(*ConveyorIO70150.xPosLimit:=X49;*)						
ConveyorIO70150.xCWPresent:=X48;						
Y248:=ConveyorIO70150.xMotorCW;						
ConveyorIO70150.xForward:=M564;						
M350:= NOT ConveyorIO70150.xEmpty;						
M749:=ConveyorIO70150.xError;						
ConveyorIO70150.diDeviceID:=70150;						

ConveyorIO70151.xPosLimit:=X4B;						
ConveyorIO70151.xCWPresent:=X4A;						
Y249:=ConveyorIO70151.xMotorCCW;						
ConveyorIO70151.xBackward:=M565;						
M351:= NOT ConveyorIO70151.xEmpty;						
M750:=ConveyorIO70151.xError;						
ConveyorIO70151.diDeviceID:=70151;						

ConveyorIO70152.xCWPresent:=X4D;						
Y24A:=ConveyorIO70152.xMotorCW;						
ConveyorIO70152.xForward:=M566;						
M352:= NOT ConveyorIO70152.xEmpty;						
M751:=ConveyorIO70152.xError;						
ConveyorIO70152.diDeviceID:=70152;			
ConveyorIO70152.tLoadDelay:=T#7S;			

ConveyorIO70153.xCWPresent:=X4D;						
Y24B:=ConveyorIO70153.xMotorCW;						
ConveyorIO70153.xForward:=M567;						
M353:= NOT ConveyorIO70153.xEmpty;						
M752:=ConveyorIO70153.xError;						
ConveyorIO70153.diDeviceID:=70153;						

ConveyorIO70154.xPosLimit:=X4F;						
ConveyorIO70154.xCWPresent:=X4E;						
Y24C:=ConveyorIO70154.xMotorCW;						
ConveyorIO70154.xForward:=M568;						
M354:= NOT ConveyorIO70154.xEmpty;						
M753:=ConveyorIO70154.xError;						
ConveyorIO70154.diDeviceID:=70154;		
ConveyorIO70154.tLoadDelay:=T#4S;				
				
ConveyorIO70155.xCWPresent:=X50;						
Y24D:=ConveyorIO70155.xMotorCW;						
ConveyorIO70155.xBackward:=M569;						
M355:= NOT ConveyorIO70155.xEmpty;						
M754:=ConveyorIO70155.xError;						
ConveyorIO70155.diDeviceID:=70155;		
ConveyorIO70155.tLoadDelay:=T#4S;						

ConveyorIO70156.xPosLimit:=NOT  X53;						
ConveyorIO70156.xCWPresent:=X52;						
Y24E:=ConveyorIO70156.xMotorCW;						
ConveyorIO70156.xForward:=M570;						
M356:= NOT ConveyorIO70156.xEmpty;						
M755:=ConveyorIO70156.xError;						
ConveyorIO70156.diDeviceID:=70156;						

ConveyorIO70157.xCWPresent:=X54;						
Y24F:=ConveyorIO70157.xMotorCW;						
ConveyorIO70157.xForward:=M571;						
M357:= NOT ConveyorIO70157.xEmpty;						
M756:=ConveyorIO70157.xError;						
ConveyorIO70157.diDeviceID:=70157;						

ConveyorIO70158.xPosLimit:=X56;						
ConveyorIO70158.xCWPresent:=X55;						
Y250:=ConveyorIO70158.xMotorCW;						
ConveyorIO70158.xForward:=M572;						
M358:= NOT ConveyorIO70158.xEmpty;						
M757:=ConveyorIO70158.xError;						
ConveyorIO70158.diDeviceID:=70158;						

(*ConveyorIO70159.xPosLimit:=X57;	*)					
ConveyorIO70159.xCWPresent:=X57;						
Y251:=ConveyorIO70159.xMotorCW;						
ConveyorIO70159.xBackward:=M573;						
M359:= NOT ConveyorIO70159.xEmpty;						
M758:=ConveyorIO70159.xError;						
ConveyorIO70159.diDeviceID:=70159;						

ConveyorIO70160.xCWPresent:=X59;						
Y252:=ConveyorIO70160.xMotorCW;						
ConveyorIO70160.xForward:=M574;						
M360:= NOT ConveyorIO70160.xEmpty;						
M759:=ConveyorIO70160.xError;						
ConveyorIO70160.diDeviceID:=70160;		
ConveyorIO70160.tLoadDelay:=T#7S;				

ConveyorIO70161.xCWPresent:=X5A;						
Y253:=ConveyorIO70161.xMotorCW;						
ConveyorIO70161.xForward:=M575;						
M361:= NOT ConveyorIO70161.xEmpty;						
M760:=ConveyorIO70161.xError;						
ConveyorIO70161.diDeviceID:=70161;						

(*ConveyorIO70162.xPosLimit:=X5C;	*)					
ConveyorIO70162.xCWPresent:=X5B;						
Y254:=ConveyorIO70162.xMotorCW;						
ConveyorIO70162.xForward:=M576;						
M362:= NOT ConveyorIO70162.xEmpty;						
M761:=ConveyorIO70162.xError;						
ConveyorIO70162.diDeviceID:=70162;						
ConveyorIO70162.tLoadDelay:=T#5S;

(*ConveyorIO70163.xPosLimit:=X5E;	*)					
ConveyorIO70163.xCWPresent:=X5D;						
Y305:=ConveyorIO70163.xMotorCW ;						
ConveyorIO70163.xBackward:=M577;						
M363:= NOT ConveyorIO70163.xEmpty;						
M762:=ConveyorIO70163.xError;						
ConveyorIO70163.diDeviceID:=70163;	
ConveyorIO70163.tLoadDelay:=t#4s;

ConveyorIO70164.xCWPresent:=X5F;						
Y256:=ConveyorIO70164.xMotorCW OR M800;						
ConveyorIO70164.xForward:=M578;						
M364:= NOT ConveyorIO70164.xEmpty;						
M763:=ConveyorIO70164.xError;						
ConveyorIO70164.diDeviceID:=70164;			
ConveyorIO70164.tLoadDelay:=T#4s;			

ConveyorIO70165.xCWPresent:=X61;						
Y257:=ConveyorIO70165.xMotorCW OR ConveyorIO70165_2.xMotorCW;						
ConveyorIO70165.xForward:=M579;						
M365:= NOT ConveyorIO70165.xEmpty;						
M764:=ConveyorIO70165.xError;						
ConveyorIO70165.diDeviceID:=70165;		
ConveyorIO70165.tLoadDelay:=T#4200MS;


ConveyorIO70165_1.xCWPresent:=	X5F;
ConveyorIO70165_1.diDeviceID:=70164;		

ConveyorIO70165_2.xCWPresent:=	X60;
ConveyorIO70165_2.diDeviceID:=70165;		
ConveyorIO70165_2.tLoadDelay:=T#4500MS;

ConveyorIO70166.xCWPresent:=X62;						
Y258:=ConveyorIO70166.xMotorCW;						
ConveyorIO70166.xForward:=M580;						
M366:= NOT ConveyorIO70166.xEmpty;						
M765:=ConveyorIO70166.xError;						
ConveyorIO70166.diDeviceID:=70166;						
ConveyorIO70166.tLoadDelay:=T#6S;

ConveyorIO70167.xCWPresent:=X63;						
Y259:=ConveyorIO70167.xMotorCW;						
ConveyorIO70167.xForward:=M581;						
M367:= NOT ConveyorIO70167.xEmpty;						
M766:=ConveyorIO70167.xError;						
ConveyorIO70167.diDeviceID:=70167;		
ConveyorIO70167.tLoadDelay:=T#8S;				

ConveyorIO70168.xCWPresent:=X65;						
Y25A:=ConveyorIO70168.xMotorCW OR ConveyorIO70168_1.xMotorCW;						
ConveyorIO70168.xForward:=M582;						
M368:= NOT ConveyorIO70168.xEmpty;						
M767:=ConveyorIO70168.xError;						
ConveyorIO70168.diDeviceID:=70168;		
ConveyorIO70168.tLoadDelay:=T#6S;

ConveyorIO70168_1.xCWPresent:=X64;
ConveyorIO70168_1.diDeviceID:=70168;	
ConveyorIO70168_1.tLoadDelay:=T#6S;

ConveyorIO70169.xCWPresent:=X64;						
ConveyorIO70169.xCCWPresent:=X65;						
Y25B:=ConveyorIO70169.xMotorCW;						
ConveyorIO70169.xForward:=M583;						
M369:= NOT ConveyorIO70169.xEmpty;						
M768:=ConveyorIO70169.xError;						
ConveyorIO70169.diDeviceID:=70169;						

(*ConveyorIO70170.xPosLimit:=X67;	*)					
ConveyorIO70170.xCWPresent:=X65;						
Y25C:=ConveyorIO70170.xMotorCW;						
ConveyorIO70170.xForward:=M584;						
M370:= NOT ConveyorIO70170.xEmpty;						
M769:=ConveyorIO70170.xError;						
ConveyorIO70170.diDeviceID:=70170;						

ConveyorIO70171.xCWPresent:=X68 OR X61;
ConveyorIO70171.xCcWPresent:=X68 OR X61;
Y25D:=ConveyorIO70171.xMotorCW;						
Y25E:=ConveyorIO70171.xMotorCCW;						
ConveyorIO70171.xForward:=M585;						
ConveyorIO70171.xBackward:=M586;						
M371:= NOT ConveyorIO70171.xEmpty;						
M770:=ConveyorIO70171.xError;						
ConveyorIO70171.diDeviceID:=70171;		
ConveyorIO70171.tLoadDelay:=T#7s;				

ConveyorIO70172.xCcWPresent:=X62;	
ConveyorIO70172.xCWPresent:=X62;					
Y25F:=ConveyorIO70172.xMotorCW;						
Y260:=ConveyorIO70172.xMotorCCW;						
ConveyorIO70172.xForward:=M587;						
ConveyorIO70172.xBackward:=M588;						
M372:= NOT ConveyorIO70172.xEmpty;						
M771:=ConveyorIO70172.xError;						
ConveyorIO70172.diDeviceID:=70172;	
ConveyorIO70172.tLoadDelay:=t#7s;					

ConveyorIO70173.xCWPresent:=X6A;
					
Y261:=ConveyorIO70173.xMotorCW;						
Y262:=ConveyorIO70173.xMotorCCW;						
ConveyorIO70173.xForward:=M589;						
ConveyorIO70173.xBackward:=M590;						
M373:= NOT ConveyorIO70173.xEmpty;						
M772:=ConveyorIO70173.xError;						
ConveyorIO70173.diDeviceID:=70173;	
ConveyorIO70173.tLoadDelay:=t#3S;					

ConveyorIO70173_1.xCWPresent:=X63;
ConveyorIO70173_1.diDeviceID:=70173;
ConveyorIO70173_1.tLoadDelay:=T#5S;

ConveyorIO70174.xCWPresent:=X6B;						
Y263:=ConveyorIO70174.xMotorCW;						
ConveyorIO70174.xForward:=M591;						
M374:= NOT ConveyorIO70174.xEmpty;						
M773:=ConveyorIO70174.xError;						
ConveyorIO70174.diDeviceID:=70174;						
ConveyorIO70174.tLoadDelay:=T#5S;

(*ConveyorIO70175.xPosLimit:=X6D;*)						
ConveyorIO70175.xCWPresent:=X70;						
Y264:=ConveyorIO70175.xMotorCW OR ConveyorIO70175_2.xMotorCW ;						
ConveyorIO70175.xForward:=M592;						
M375:= NOT ConveyorIO70175.xEmpty;						
M774:=ConveyorIO70175.xError;						
ConveyorIO70175.diDeviceID:=70175;		
ConveyorIO70175.tLoadDelay:=T#4000MS;


ConveyorIO70175_1.xCWPresent:=	X6B;
ConveyorIO70175_1.diDeviceID:=70174;			

ConveyorIO70175_2.xCWPresent:=	X6C;
ConveyorIO70175_2.diDeviceID:=70175;	
ConveyorIO70175_2.tLoadDelay:=t#4500ms;

ConveyorIO70176.xCWPresent:=X71;						
Y265:=ConveyorIO70176.xMotorCW;						
ConveyorIO70176.xForward:=M593;						
M376:= NOT ConveyorIO70176.xEmpty;						
M775:=ConveyorIO70176.xError;						
ConveyorIO70176.diDeviceID:=70176;						
ConveyorIO70176.tLoadDelay:=T#6S;

ConveyorIO70177.xCWPresent:=X157 OR X72;						
Y266:=ConveyorIO70177.xMotorCW;						
ConveyorIO70177.xForward:=M594;						
M377:= NOT ConveyorIO70177.xEmpty;						
M776:=ConveyorIO70177.xError;						
ConveyorIO70177.diDeviceID:=70177;		
ConveyorIO70177.tLoadDelay:=T#5S;				

ConveyorIO70178.xCWPresent:=X73;						
Y267:=ConveyorIO70178.xMotorCW;						
ConveyorIO70178.xForward:=M595;						
M378:= NOT ConveyorIO70178.xEmpty;						
M777:=ConveyorIO70178.xError;						
ConveyorIO70178.diDeviceID:=70178;		
ConveyorIO70178.tLoadDelay:=T#1S;				

ConveyorIO70179.xCWPresent:=X74;						
Y268:=ConveyorIO70179.xMotorCW;						
ConveyorIO70179.xForward:=M596;						
M379:= NOT ConveyorIO70179.xEmpty;						
M778:=ConveyorIO70179.xError;						
ConveyorIO70179.diDeviceID:=70179;						

ConveyorIO70180.xCWPresent:=X75;						
Y269:=ConveyorIO70180.xMotorCW;						
ConveyorIO70180.xForward:=M597;						
M380:= NOT ConveyorIO70180.xEmpty;						
M779:=ConveyorIO70180.xError;						
ConveyorIO70180.diDeviceID:=70180;	
ConveyorIO70180.tLoadDelay:=T#4S;					

ConveyorIO70181.xPosLimit:=NOT XBD;
ConveyorIO70181.xCWPresent:=XF0;						
Y26A:=ConveyorIO70181.xMotorCW;						
ConveyorIO70181.xForward:=M598;						
M381:= NOT ConveyorIO70181.xEmpty;						
M780:=ConveyorIO70181.xError;						
ConveyorIO70181.diDeviceID:=70181;						

ConveyorIO70182.xCWPresent:=X70;						
Y26B:=ConveyorIO70182.xMotorCW;						
Y26C:=ConveyorIO70182.xMotorCCW;						
ConveyorIO70182.xForward:=M599;						
ConveyorIO70182.xBackward:=M600;						
M382:= NOT ConveyorIO70182.xEmpty;						
M781:=ConveyorIO70182.xError;						
ConveyorIO70182.diDeviceID:=70182;
ConveyorIO70182.tLoadDelay:=T#5S;						

ConveyorIO70183.xCWPresent:=X71;						
Y26D:=ConveyorIO70183.xMotorCW;						
Y26E:=ConveyorIO70183.xMotorCCW;						
ConveyorIO70183.xForward:=M601;						
ConveyorIO70183.xBackward:=M602;						
M383:= NOT ConveyorIO70183.xEmpty;						
M782:=ConveyorIO70183.xError;						
ConveyorIO70183.diDeviceID:=70183;				
ConveyorIO70183.tLoadDelay:=T#6S;		

ConveyorIO70184.xCWPresent:=X78;						
Y26F:=ConveyorIO70184.xMotorCW;						
Y270:=ConveyorIO70184.xMotorCCW;						
ConveyorIO70184.xForward:=M603;						
ConveyorIO70184.xBackward:=M604;						
M384:= NOT ConveyorIO70184.xEmpty;						
M783:=ConveyorIO70184.xError;						
ConveyorIO70184.diDeviceID:=70184;						

ConveyorIO70184_1.xCWPresent:=X72;
ConveyorIO70184_1.diDeviceID:=70184;
ConveyorIO70184_1.tLoadDelay:=T#5S;

ConveyorIO70185.xCWPresent:=X79;						
Y271:=ConveyorIO70185.xMotorCW;						
ConveyorIO70185.xForward:=M605;						
M385:= NOT ConveyorIO70185.xEmpty;						
M784:=ConveyorIO70185.xError;						
ConveyorIO70185.diDeviceID:=70185;	

ConveyorIO70190.xCWPresent:=X3F;						
Y2FA:=ConveyorIO70190.xMotorCCW;	
Y2FB:=ConveyorIO70190.xMotorCW;					
ConveyorIO70190.xForward:=M612;	
ConveyorIO70190.xBackward:=M622;					
(*M385:= NOT ConveyorIO70185.xEmpty;						
M784:=ConveyorIO70185.xError;	*)					
ConveyorIO70190.diDeviceID:=70190;	

ConveyorIO70191.xCWPresent:=X134;
ConveyorIO70191.xCCWPresent:=X134;
Y2FC:=ConveyorIO70191.xMotorCW;
Y2FD:=ConveyorIO70191.xMotorCCW;
ConveyorIO70191.xForward:=M623;
ConveyorIO70191.xBackward:=M624;
ConveyorIO70191.diDeviceID:=70191;
ConveyorIO70191.tLoadDelay:=t#10s;

ConveyorIO70192.xCWPresent:=X4D;
Y2FE:=ConveyorIO70192.xMotorCW;
Y2FF:=ConveyorIO70192.xMotorCCW;
ConveyorIO70192.xForward:=M623;
ConveyorIO70192.xBackward:=M624;
ConveyorIO70192.diDeviceID:=70192;


ConveyorIO70193.xCWPresent:=X136;						
ConveyorIO70193.xCCWPresent:=X136;						
Y300:=ConveyorIO70193.xMotorCW;		
Y301:=ConveyorIO70193.xMotorCCW;					
ConveyorIO70193.xForward:=M678;						
(*M385:= NOT ConveyorIO70185.xEmpty;						
M784:=ConveyorIO70185.xError;	*)					
ConveyorIO70193.diDeviceID:=70193;	
ConveyorIO70193.tLoadDelay:=T#10s;	

ConveyorIO70194.xCWPresent:=X59;						
Y302:=ConveyorIO70194.xMotorCW;		
Y303:=ConveyorIO70194.xMotorCCW;					
ConveyorIO70194.xForward:=M678;						
(*M385:= NOT ConveyorIO70185.xEmpty;						
M784:=ConveyorIO70185.xError;	*)					
ConveyorIO70194.diDeviceID:=70194;	
ConveyorIO70194.tLoadDelay:=T#5s;	

ConveyorIO70195.xCWPresent:=X138;						
Y2EC:=ConveyorIO70195.xMotorCW;						
ConveyorIO70195.xForward:=M611;						
(*M385:= NOT ConveyorIO70185.xEmpty;						
M784:=ConveyorIO70185.xError;	*)					
ConveyorIO70195.diDeviceID:=70195;	
ConveyorIO70195.tLoadDelay:=T#4s;	

ConveyorIO70196.xCWPresent:=X139;						
Y2ED:=ConveyorIO70196.xMotorCW;						
ConveyorIO70196.xForward:=M613;						
(*M385:= NOT ConveyorIO70185.xEmpty;						
M784:=ConveyorIO70185.xError;	*)					
ConveyorIO70196.diDeviceID:=70196;	
ConveyorIO70196.tLoadDelay:=t#4s;		

ConveyorIo70197.xCWPresent:=X13A;
Y2EE:=ConveyorIo70197.xMotorCW;
ConveyorIO70197.xForward:=M625;
ConveyorIo70197.diDeviceID:=70197;
ConveyorIo70197.tLoadDelay:=T#2s;

ConveyorIO70198.xCWPresent:=X13B;
Y2EF:=ConveyorIO70198.xMotorCW;
ConveyorIO70198.xForward:=M626;
ConveyorIO70198.diDeviceID:=70198;		

ConveyorIO70199.xCWPresent:=X13C;
Y2F0:=ConveyorIO70199.xMotorCW;
ConveyorIO70199.xForward:=M626;
ConveyorIO70199.diDeviceID:=70199;		

ConveyorIO701100.xCWPresent:=X13D;
Y2F1:=ConveyorIO701100.xMotorCW;
ConveyorIO701100.xForward:=M626;
ConveyorIO701100.diDeviceID:=701100;		
ConveyorIO701100.tLoadDelay:=t#3S;

ConveyorIO701102.xCWPresent:=X13F;
Y2F3:=ConveyorIO701102.xMotorCW ;
ConveyorIO701102.xForward:=M679;
ConveyorIO701102.diDeviceID:=701103;
ConveyorIO701102.tLoadDelay:=T#2s;

ConveyorIO701103.xCWPresent:=X140;
Y304:=ConveyorIO701103.xMotorCW ;
ConveyorIO701103.xForward:=M679;
ConveyorIO701103.diDeviceID:=701103;
ConveyorIO701103.tLoadDelay:=T#4s;

ConveyorIO701104.xCWPresent:=X141;
Y255:=ConveyorIO701104.xMotorCW ;
ConveyorIO701104.diDeviceID:=701104;
ConveyorIO701104.tLoadDelay:=T#4s;

ConveyorIO701111.xCWPresent:=X148;
ConveyorIO701111.xPosLimit:=NOT X150;
Y306:=ConveyorIO701111.xMotorCW OR ConveyorIO701111_1.xMotorCW ;
ConveyorIO701111.xForward:=	M614;
ConveyorIO701111.diDeviceID:=701111;

ConveyorIO701111_1.xCWPresent:=X14A;
ConveyorIO701111_1.diDeviceID:=701111;

ConveyorIO701113.xCWPresent:=X14A;
Y308:=ConveyorIO701113.xMotorCW ;
ConveyorIO701113.xForward:=M615;
ConveyorIO701113.diDeviceID:=701113;
ConveyorIO701113.tLoadDelay:=T#5s;

ConveyorIO701114.xCWPresent:=X15B;
Y309:=ConveyorIO701114.xMotorCW;
ConveyorIO701114.xForward:=M616;
ConveyorIO701114.diDeviceID:=701114;
ConveyorIO701114.tLoadDelay:=T#2S;

ConveyorIO701115.xCWPresent:=X14B;
Y30A:=ConveyorIO701115.xMotorCW;
ConveyorIO701115.xForward:=M617;
ConveyorIO701115.diDeviceID:=701115;
		
					
Switch70301(ConveyorEntryIO:= ConveyorIO70104 ,ConveyorExitIO:=ConveyorIO70105 ,SwitchIO:=SwitchIO70301 );
SwitchIO70301.xLiftCylinderExtendButton:=M606;
SwitchIO70301.xLiftCylinderRetractButton:=M607;
SwitchIO70301.xLiftCylinderExtendDetect:=XBF;
SwitchIO70301.xLiftCylinderRetractDetect:=XBE;
Y2AA:=SwitchIO70301.xLiftCylinderExtend;

Switch70312(ConveyorEntryIO:= ConveyorIO70191 ,ConveyorExitIO:= ConveyorIO70148_1,SwitchIO:=SwitchIO70312);
SwitchIO70312.xLiftCylinderExtendButton:=M635;
SwitchIO70312.xLiftCylinderRetractButton:=M636;
SwitchIO70312.xLiftCylinderExtendDetect:=XD4;
SwitchIO70312.xLiftCylinderRetractDetect:=XD5;
Y2C0:=SwitchIO70312.xLiftCylinderExtend;

(*Switch70316(ConveyorEntryIO:= ConveyorIO70164 ,ConveyorExitIO:= ConveyorIO70165_1 ,SwitchIO:= SwitchIO70316 );
SwitchIO70316.xLiftCylinderExtendButton:=M627;
SwitchIO70316.xLiftCylinderRetractButton:=M628;
SwitchIO70316.xLiftCylinderExtendDetect:=XDC;
SwitchIO70316.xLiftCylinderRetractDetect:=XDD;
Y2C8:=SwitchIO70316.xLiftCylinderExtend;*)

(*IF m_xOCV2_1UnloadRequest THEN *)(*有OCV2下料请求的时候顶升移载反向*)
	(*Switch70317(ConveyorEntryIO:= ConveyorIO70171  ,ConveyorExitIO:=ConveyorIO70165  ,SwitchIO:= SwitchIO70317);
	SwitchIO70317.xLiftCylinderExtendInit:=0;
	ConveyorIO70171.xloadCCW:=1;*)(*入料线体上料方向反向*)
(*	ELSE
	Switch70317(ConveyorEntryIO:= ConveyorIO70165  ,ConveyorExitIO:= ConveyorIO70171 ,SwitchIO:= SwitchIO70317);
	SwitchIO70317.xLiftCylinderExtendInit:=1;
END_IF;
SwitchIO70317.xLiftCylinderExtendButton:=M629;
SwitchIO70317.xLiftCylinderRetractButton:=M630;
SwitchIO70317.xLiftCylinderExtendDetect:=XDE;
SwitchIO70317.xLiftCylinderRetractDetect:=XDF;
Y2CA:=SwitchIO70317.xLiftCylinderExtend;*)

(*IF m_xOCV2_2UnloadRequest THEN 
	Switch70318(ConveyorEntryIO:= ConveyorIO70172  ,ConveyorExitIO:=ConveyorIO70166  ,SwitchIO:=SwitchIO70318);
	SwitchIO70318.xLiftCylinderExtendInit:=0;
	ConveyorIO70172.xloadCCW:=1;
	ELSE
	Switch70318(ConveyorEntryIO:= ConveyorIO70166  ,ConveyorExitIO:= ConveyorIO70172 ,SwitchIO:= SwitchIO70318);
	SwitchIO70318.xLiftCylinderExtendInit:=1;
END_IF;
SwitchIO70318.xLiftCylinderExtendButton:=M631;
SwitchIO70318.xLiftCylinderRetractButton:=M632;
SwitchIO70318.xLiftCylinderExtendDetect:=XE0;
SwitchIO70318.xLiftCylinderRetractDetect:=XE1;
Y2CC:=SwitchIO70318.xLiftCylinderExtend;*)


Switch70326(ConveyorEntryIO:= ConveyorIO701113 ,ConveyorExitIO:= ConveyorIO701111_1 ,SwitchIO:= SwitchIO70326);
SwitchIO70326.xLiftCylinderExtendButton:=M618;
SwitchIO70326.xLiftCylinderRetractButton:=M619;
SwitchIO70326.xLiftCylinderExtendDetect:=X153;
SwitchIO70326.xLiftCylinderRetractDetect:=X154;
Y2DC:=SwitchIO70326.xLiftCylinderExtend;

Switch70311(ConveyorEntryIO:= ConveyorIO70144 ,ConveyorExitIO:= ConveyorIO70190 ,SwitchIO:=SwitchIO70311 );
SwitchIO70311.xLiftCylinderExtendButton:=M620;
SwitchIO70311.xLiftCylinderRetractButton:=M621;
SwitchIO70311.xLiftCylinderExtendDetect:=XD2;
SwitchIO70311.xLiftCylinderRetractDetect:=XD3;
Y2BE:=SwitchIO70311.xLiftCylinderExtend;
SwitchIo70311.xLiftCylinderExtendInit:=1;

Switch70319(ConveyorEntryIO:= ConveyorIO70167 ,ConveyorExitIO:=ConveyorIO70173 ,SwitchIO:= SwitchIO70319 );
SwitchIO70319.xLiftCylinderExtendButton:=M633;
SwitchIO70319.xLiftCylinderRetractButton:=M634;
SwitchIO70319.xLiftCylinderExtendDetect:=XE2;
SwitchIO70319.xLiftCylinderRetractDetect:=XE3;
(*Y2CE:=SwitchIO70319.xLiftCylinderExtend;*)
SwitchIO70319.xLiftCylinderExtendInit:=1;

(*Switch70320(ConveyorEntryIO:= ConveyorIO70169 ,ConveyorExitIO:= ConveyorIO70170 ,SwitchIO:= SwitchIO70320 );
SwitchIO70320.xLiftCylinderExtendButton:=M635;
SwitchIO70320.xLiftCylinderRetractButton:=M636;
SwitchIO70320.xLiftCylinderExtendDetect:=XE4;
SwitchIO70320.xLiftCylinderRetractDetect:=XE5;
Y2D0:=SwitchIO70320.xLiftCylinderExtend;
SwitchIO70320.xLiftCylinderExtendInit:=1;*)

Lift70207(ShuttleCarInOut:= LifterIO70207 );
LifterIO70207.xArrive:= ShuttleCarCurrentPosition( LifterIO70207.xPresentDetect1 OR LifterIO70207.xPresentDetect2 ,
																						 LifterIO70207.xPresentDetect1 , 
																						 LifterIO70207.xPresentDetect2 , 
																						 FALSE , 
																						 LifterIO70207.iCurrentPos );
LifterIO70207.xForward:=M608;
LifterIO70207.xBackward:=M609;
LifterIO70207.xCylinder:=1;
Y29C:=LifterIO70207.xCW;
Y29D:=LifterIO70207.xCCW;
LifterIO70207.xPresentDetect1:=XB0;
LifterIO70207.xPresentDetect2:=XB1;
LifterIO70207.tSetOverTime:=T#30s;

Lift70208(ShuttleCarInOut:= LifterIO70208 );
LifterIO70208.xArrive:= ShuttleCarCurrentPosition( LifterIO70208.xPresentDetect1 OR LifterIO70208.xPresentDetect2 ,
																						 LifterIO70208.xPresentDetect1 , 
																						 LifterIO70208.xPresentDetect2 , 
																						 FALSE , 
																						 LifterIO70208.iCurrentPos );
LifterIO70208.xForward:=M629;
LifterIO70208.xBackward:=M630;
LifterIO70208.xCylinder:=1;
Y29E:=LifterIO70208.xCW;
Y29F:=LifterIO70208.xCCW;
LifterIO70208.xPresentDetect1:=XB2;
LifterIO70208.xPresentDetect2:=XB3;
LifterIO70208.tSetOverTime:=T#30s;

Folder70201(FolderIO:= FolderIO70201 ,FolderConveyorIO:= ConveyorIO70140 ,i_xAuto:=m_xFolder70201Atuo ,i_xManual:= NOT m_xFolder70201Atuo );(*静置入口叠盘*)
FolderIO70201.i_xCylinderDownExtendButton:=M637;
FolderIO70201.i_xCylinderDownExtendDetect:=X83;
FolderIO70201.i_xCylinderDownRetractButton:=M638;
FolderIO70201.i_xCylinderDownRetractDetect:=X82;
FolderIO70201.i_xCylinderGrabExtendButton:=M639;
FolderIO70201.i_xCylinderGrabExtendDetect:=X86;
FolderIO70201.i_xCylinderGrabRetractButton:=M640;
FolderIO70201.i_xCylinderGrabRetractDetect:=X87;
FolderIO70201.i_xCylinderUpExtendButton:=M641;
FolderIO70201.i_xCylinderUpExtendDetect:=X81;
FolderIO70201.i_xCylinderUpRetractButton:=M642;
FolderIO70201.i_xCylinderUpRetractDetect:=X80;
Y278:=FolderIO70201.o_xCylinderDownExtend;
Y279:=FolderIO70201.o_xCylinderDownRetract;
Y27D:=FolderIO70201.o_xCylinderGrabExtend;
Y27C:=FolderIO70201.o_xCylinderGrabRetract;
Y27A:=FolderIO70201.o_xCylinderUpExtend;
Y27B:=FolderIO70201.o_xCylinderUpRetract;

DivideFolder70204(FolderIO:=DivideFolderIO70204 ,FolderConveyorIO:=ConveyorIO70165_2,i_xAuto:= m_xDivideFolder70204Auto);(*OCV2入口拆盘*)
DivideFolderIO70204.i_xCylinderDownExtendButton:=M644;
DivideFolderIO70204.i_xCylinderDownRetractButton:=M645;
DivideFolderIO70204.i_xCylinderGrabExtendButton:=M646;
DivideFolderIO70204.i_xCylinderGrabRetractButton:=M647;
DivideFolderIO70204.i_xCylinderUpExtendButton:=M648;
DivideFolderIO70204.i_xCylinderUpRetractButton:=M649;
DivideFolderIO70204.i_xCylinderDownExtendDetect:=X98;
DivideFolderIO70204.i_xCylinderDownRetractDetect:=X99;
DivideFolderIO70204.i_xCylinderGrabExtendDetect:=X9E;
DivideFolderIO70204.i_xCylinderGrabRetractDetect:=X9F;
DivideFolderIO70204.i_xCylinderUpExtendDetect:=X9A;
DivideFolderIO70204.i_xCylinderUpRetractDetect:=X9B;
DivideFolderIO70204.i_xTrayDetect:=X27;
Y28A:=DivideFolderIO70204.o_xCylinderDownExtend;
Y28D:=DivideFolderIO70204.o_xCylinderDownRetract;
Y28F:=DivideFolderIO70204.o_xCylinderGrabExtend;
Y28E:=DivideFolderIO70204.o_xCylinderGrabRetract;
Y28C:=DivideFolderIO70204.o_xCylinderUpExtend;
Y28B:=DivideFolderIO70204.o_xCylinderUpRetract;

Folder70205(FolderIO:= FolderIO70205 ,FolderConveyorIO:= ConveyorIO70168_1 ,i_xAuto:=m_xFolder70205Atuo ,i_xManual:= NOT m_xFolder70205Atuo );(*OCV2出口叠盘*)
FolderIO70205 .i_xCylinderDownExtendButton:=M650;
FolderIO70205 .i_xCylinderDownExtendDetect:=XA2;
FolderIO70205 .i_xCylinderDownRetractButton:=M651;
FolderIO70205 .i_xCylinderDownRetractDetect:=XA3;
FolderIO70205 .i_xCylinderGrabExtendButton:=M652;
FolderIO70205 .i_xCylinderGrabExtendDetect:=XA6;
FolderIO70205 .i_xCylinderGrabRetractButton:=M653;
FolderIO70205 .i_xCylinderGrabRetractDetect:=XA7;
FolderIO70205 .i_xCylinderUpExtendButton:=M654;
FolderIO70205 .i_xCylinderUpExtendDetect:=XA0;
FolderIO70205 .i_xCylinderUpRetractButton:=M655;
FolderIO70205 .i_xCylinderUpRetractDetect:=XA1;
FolderIO70205 .i_xTrayDetect:=XFD;
Y291:=FolderIO70205 .o_xCylinderDownExtend;
Y293:=FolderIO70205 .o_xCylinderDownRetract;
Y294:=FolderIO70205 .o_xCylinderGrabExtend;
Y295:=FolderIO70205 .o_xCylinderGrabRetract;
Y290:=FolderIO70205 .o_xCylinderUpExtend;
Y292:=FolderIO70205 .o_xCylinderUpRetract;


DivideFolder70206(FolderIO:= DivideFolderIO70206 ,FolderConveyorIO:=ConveyorIO70175_2,i_xAuto:= m_xDivideFolder70206Auto );(*OCV3入口拆盘*)
DivideFolderIO70206 .i_xCylinderDownExtendButton:=M657;
DivideFolderIO70206 .i_xCylinderDownRetractButton:=M658;
DivideFolderIO70206 .i_xCylinderGrabExtendButton:=M659;
DivideFolderIO70206 .i_xCylinderGrabRetractButton:=M660;
DivideFolderIO70206 .i_xCylinderUpExtendButton:=M661;
DivideFolderIO70206 .i_xCylinderUpRetractButton:=M662;
DivideFolderIO70206 .i_xCylinderDownExtendDetect:=XAA;
DivideFolderIO70206 .i_xCylinderDownRetractDetect:=XAB;
DivideFolderIO70206 .i_xCylinderGrabExtendDetect:=XAC;
DivideFolderIO70206 .i_xCylinderGrabRetractDetect:=XAD;
DivideFolderIO70206 .i_xCylinderUpExtendDetect:=XA9;
DivideFolderIO70206 .i_xCylinderUpRetractDetect:=XA8;
DivideFolderIO70206 .i_xTrayDetect:=XE6;
Y297:=DivideFolderIO70206 .o_xCylinderDownExtend;
Y298:=DivideFolderIO70206 .o_xCylinderDownRetract;
Y29A:=DivideFolderIO70206 .o_xCylinderGrabExtend;
Y29B:=DivideFolderIO70206 .o_xCylinderGrabRetract;
Y296:=DivideFolderIO70206 .o_xCylinderUpExtend;
Y299:=DivideFolderIO70206 .o_xCylinderUpRetract;



(*与上位机通讯程序*)
ComConveyor70104(ConveyorIO:= ConveyorIO70140_1,CommunicationIO:= ComConveyorIO70104);
ComConveyor70106(ConveyorIO:= ConveyorIO70140,CommunicationIO:= ComConveyorIO70106);(*线体更改*)
ComConveyor70144(ConveyorIO:= ConveyorIO70144,CommunicationIO:= ComConveyorIO70144);
ComConveyor70152(ConveyorIO:= ConveyorIO70152,CommunicationIO:= ComConveyorIO70152);
ComConveyor70146(ConveyorIO:= ConveyorIO70146,CommunicationIO:= ComConveyorIO70146);
ComConveyor70195(ConveyorIO:= ConveyorIO70195,CommunicationIO:= ComConveyorIO70195);
ComConveyor70147(ConveyorIO:= ConveyorIO70147,CommunicationIO:= ComConveyorIO70147);
ComConveyor70196(ConveyorIO:= ConveyorIO70196,CommunicationIO:= ComConveyorIO70196);
ComConveyor70154(ConveyorIO:= ConveyorIO70154,CommunicationIO:= ComConveyorIO70154);
ComConveyor70199(ConveyorIO:= ConveyorIO70199,CommunicationIO:= ComConveyorIO70199);
ComConveyor70155(ConveyorIO:= ConveyorIO70155,CommunicationIO:= ComConveyorIO70155);
ComConveyor701100(ConveyorIO:= ConveyorIO701100,CommunicationIO:= ComConveyorIO701100);
ComConveyor701115(ConveyorIO:= ConveyorIO701115,CommunicationIO:= ComConveyorIO701115);
ComConveyor701114(ConveyorIO:= ConveyorIO701114,CommunicationIO:= ComConveyorIO701114);
ComConveyor70197(ConveyorIO:= ConveyorIO70197,CommunicationIO:= ComConveyorIO70197);
ComConveyor70150(ConveyorIO:= ConveyorIO70150,CommunicationIO:= ComConveyorIO70150);
ComConveyor70151(ConveyorIO:= ConveyorIO70151,CommunicationIO:= ComConveyorIO70151);
ComConveyor70198(ConveyorIO:= ConveyorIO70198,CommunicationIO:= ComConveyorIO70198);
ComConveyor701101(ConveyorIO:= ConveyorIO701101,CommunicationIO:= ComConveyorIO701101);
ComConveyor70158(ConveyorIO:= ConveyorIO70158,CommunicationIO:= ComConveyorIO70158);
ComConveyor701111(ConveyorIO:= ConveyorIO701111,CommunicationIO:= ComConveyorIO701111);
ComConveyor70148(ConveyorIO:= ConveyorIO70148,CommunicationIO:= ComConveyorIO70148);
ComConveyor70156(ConveyorIO:= ConveyorIO70156,CommunicationIO:= ComConveyorIO70156);
ComConveyor701116(ConveyorIO:= ConveyorIO701116,CommunicationIO:= ComConveyorIO701116);
ComConveyor70164(ConveyorIO:= ConveyorIO70164,CommunicationIO:= ComConveyorIO70164);
ComConveyor70174(ConveyorIO:= ConveyorIO70174,CommunicationIO:= ComConveyorIO70174);
ComConveyor70169(ConveyorIO:= ConveyorIO70169,CommunicationIO:= ComConveyorIO70169);
ComConveyor70170(ConveyorIO:= ConveyorIO70170,CommunicationIO:= ComConveyorIO70170);
ComConveyor70160(ConveyorIO:= ConveyorIO70160,CommunicationIO:= ComConveyorIO70160);
ComConveyor70162(ConveyorIO:= ConveyorIO70162,CommunicationIO:= ComConveyorIO70162);
ComConveyor701103(ConveyorIO:= ConveyorIO701103,CommunicationIO:= ComConveyorIO701103);
ComConveyor70163(ConveyorIO:= ConveyorIO70163,CommunicationIO:= ComConveyorIO70163);
ComConveyor701104(ConveyorIO:= ConveyorIO701104,CommunicationIO:= ComConveyorIO701104);
ComConveyor701102(ConveyorIO:= ConveyorIO701102,CommunicationIO:= ComConveyorIO701102);
ComConveyor70159(ConveyorIO:= ConveyorIO70159,CommunicationIO:= ComConveyorIO70159);
ComConveyor701120(ConveyorIO:= ConveyorIO701120,CommunicationIO:= ComConveyorIO701120);
ComConveyor701119(ConveyorIO:= ConveyorIO701119,CommunicationIO:= ComConveyorIO701119);
(*ComConveyor70111(ConveyorIO:= ConveyorIO70111,CommunicationIO:= ComConveyorIO70111);
ComConveyor70112(ConveyorIO:= ConveyorIO70112,CommunicationIO:= ComConveyorIO70112);
ComConveyor701105(ConveyorIO:= ConveyorIO701105,CommunicationIO:= ComConveyorIO701105);
ComConveyor70113(ConveyorIO:= ConveyorIO70113,CommunicationIO:= ComConveyorIO70113);
ComConveyor701106(ConveyorIO:= ConveyorIO701106,CommunicationIO:= ComConveyorIO701106);
ComConveyor70114(ConveyorIO:= ConveyorIO70114,CommunicationIO:= ComConveyorIO70114);
ComConveyor70116(ConveyorIO:= ConveyorIO70116,CommunicationIO:= ComConveyorIO70116);
ComConveyor70119(ConveyorIO:= ConveyorIO70119,CommunicationIO:= ComConveyorIO70119);
ComConveyor70120(ConveyorIO:= ConveyorIO70120,CommunicationIO:= ComConveyorIO70120);
ComConveyor701107(ConveyorIO:= ConveyorIO701107,CommunicationIO:= ComConveyorIO701107);
ComConveyor70121(ConveyorIO:= ConveyorIO70121,CommunicationIO:= ComConveyorIO70121);
ComConveyor701108(ConveyorIO:= ConveyorIO701108,CommunicationIO:= ComConveyorIO701108);
ComConveyor70122(ConveyorIO:= ConveyorIO70122,CommunicationIO:= ComConveyorIO70122);
ComConveyor70124(ConveyorIO:= ConveyorIO70124,CommunicationIO:= ComConveyorIO70124);
ComConveyor70127(ConveyorIO:= ConveyorIO70127,CommunicationIO:= ComConveyorIO70127);
ComConveyor70128(ConveyorIO:= ConveyorIO70128,CommunicationIO:= ComConveyorIO70128);
ComConveyor701109(ConveyorIO:= ConveyorIO701109,CommunicationIO:= ComConveyorIO701109);
ComConveyor70129(ConveyorIO:= ConveyorIO70129,CommunicationIO:= ComConveyorIO70129);
ComConveyor701110(ConveyorIO:= ConveyorIO701110,CommunicationIO:= ComConveyorIO701110);
ComConveyor70184(ConveyorIO:= ConveyorIO70184,CommunicationIO:= ComConveyorIO70184);*)

ComConveyorIO70104.i_iResponsPCPLC:=D2000; 
ComConveyorIO70104.i_iTypeInfoPCPLC:=D2001;
ComConveyorIO70104.i_iReadWriteFlagPCPLC:=D2005; 
ComConveyorIO70104.i_iTaskProcessFlagPCPLC:=D2006; 
ComConveyorIO70104.i_iCommandPCPLC:=D2007; 
ComConveyorIO70104.i_iTaskIDPCPLC:=D2008; 
DMOV(TRUE,D2009,ComConveyorIO70104.i_diDestinationDevicePCPLC); 
ComConveyorIO70104.i_iProductIDPCPLC:=D2011;
D3000:=ComConveyorIO70104.o_iRequestPLCPC; 
D3001:=ComConveyorIO70104.o_iForceInportPLCPC;
D3002:=ComConveyorIO70104.o_iFolderNumberPLCPC;
D3003:=ComConveyorIO70104.o_iEmptyPLCPC;
D3005:=ComConveyorIO70104.o_iReadWriteFlagPLCPC; 
D3006:=ComConveyorIO70104.o_iDeviceStatusPLCPC; 
D3007:=ComConveyorIO70104.o_iTaskIDPLCPC; 
D3008:=ComConveyorIO70104.o_iProductIDPLCPC;

ComConveyorIO70106.i_iTypeInfoPCPLC:=D2031;
ComConveyorIO70106.i_iReadWriteFlagPCPLC:=D2035; 
ComConveyorIO70106.i_iTaskProcessFlagPCPLC:=D2036; 
ComConveyorIO70106.i_iCommandPCPLC:=D2037; 
ComConveyorIO70106.i_iTaskIDPCPLC:=D2038; 
DMOV(TRUE,D2039,ComConveyorIO70106.i_diDestinationDevicePCPLC); 
ComConveyorIO70106.i_iProductIDPCPLC:=D2041;
D3030:=ComConveyorIO70106.o_iRequestPLCPC; 
D3031:=ComConveyorIO70106.o_iForceInportPLCPC;
D3032:=ComConveyorIO70106.o_iFolderNumberPLCPC;
D3033:=ComConveyorIO70106.o_iEmptyPLCPC;
D3035:=ComConveyorIO70106.o_iReadWriteFlagPLCPC; 
D3036:=ComConveyorIO70106.o_iDeviceStatusPLCPC; 
D3037:=ComConveyorIO70106.o_iTaskIDPLCPC; 
D3038:=ComConveyorIO70106.o_iProductIDPLCPC;
ComConveyorIO70144.i_iResponsPCPLC:=D2045; 
ComConveyorIO70144.i_iTypeInfoPCPLC:=D2046;
ComConveyorIO70144.i_iReadWriteFlagPCPLC:=D2050; 
ComConveyorIO70144.i_iTaskProcessFlagPCPLC:=D2051; 
ComConveyorIO70144.i_iCommandPCPLC:=D2052; 
ComConveyorIO70144.i_iTaskIDPCPLC:=D2053; 
DMOV(TRUE,D2054,ComConveyorIO70144.i_diDestinationDevicePCPLC); 
ComConveyorIO70144.i_iProductIDPCPLC:=D2056;
D3045:=ComConveyorIO70144.o_iRequestPLCPC; 
D3046:=ComConveyorIO70144.o_iForceInportPLCPC;
D3047:=ComConveyorIO70144.o_iFolderNumberPLCPC;
D3048:=ComConveyorIO70144.o_iEmptyPLCPC;
D3050:=ComConveyorIO70144.o_iReadWriteFlagPLCPC; 
D3051:=ComConveyorIO70144.o_iDeviceStatusPLCPC; 
D3052:=ComConveyorIO70144.o_iTaskIDPLCPC; 
D3053:=ComConveyorIO70144.o_iProductIDPLCPC;
ComConveyorIO70152.i_iResponsPCPLC:=D2060; 
ComConveyorIO70152.i_iTypeInfoPCPLC:=D2061;
ComConveyorIO70152.i_iReadWriteFlagPCPLC:=D2065; 
ComConveyorIO70152.i_iTaskProcessFlagPCPLC:=D2066; 
ComConveyorIO70152.i_iCommandPCPLC:=D2067; 
ComConveyorIO70152.i_iTaskIDPCPLC:=D2068; 
DMOV(TRUE,D2069,ComConveyorIO70152.i_diDestinationDevicePCPLC); 
ComConveyorIO70152.i_iProductIDPCPLC:=D2071;
D3060:=ComConveyorIO70152.o_iRequestPLCPC; 
D3061:=ComConveyorIO70152.o_iForceInportPLCPC;
D3062:=ComConveyorIO70152.o_iFolderNumberPLCPC;
D3063:=ComConveyorIO70152.o_iEmptyPLCPC;
D3065:=ComConveyorIO70152.o_iReadWriteFlagPLCPC; 
D3066:=ComConveyorIO70152.o_iDeviceStatusPLCPC; 
D3067:=ComConveyorIO70152.o_iTaskIDPLCPC; 
D3068:=ComConveyorIO70152.o_iProductIDPLCPC;
ComConveyorIO70146.i_iResponsPCPLC:=D2075; 
ComConveyorIO70146.i_iTypeInfoPCPLC:=D2076;
ComConveyorIO70146.i_iReadWriteFlagPCPLC:=D2080; 
ComConveyorIO70146.i_iTaskProcessFlagPCPLC:=D2081; 
ComConveyorIO70146.i_iCommandPCPLC:=D2082; 
ComConveyorIO70146.i_iTaskIDPCPLC:=D2083; 
DMOV(TRUE,D2084,ComConveyorIO70146.i_diDestinationDevicePCPLC); 
ComConveyorIO70146.i_iProductIDPCPLC:=D2086;
D3075:=ComConveyorIO70146.o_iRequestPLCPC; 
D3076:=ComConveyorIO70146.o_iForceInportPLCPC;
D3077:=ComConveyorIO70146.o_iFolderNumberPLCPC;
D3078:=ComConveyorIO70146.o_iEmptyPLCPC;
D3080:=ComConveyorIO70146.o_iReadWriteFlagPLCPC; 
D3081:=ComConveyorIO70146.o_iDeviceStatusPLCPC; 
D3082:=ComConveyorIO70146.o_iTaskIDPLCPC; 
D3083:=ComConveyorIO70146.o_iProductIDPLCPC;
ComConveyorIO70195.i_iResponsPCPLC:=D2090; 
ComConveyorIO70195.i_iTypeInfoPCPLC:=D2091;
ComConveyorIO70195.i_iReadWriteFlagPCPLC:=D2095; 
ComConveyorIO70195.i_iTaskProcessFlagPCPLC:=D2096; 
ComConveyorIO70195.i_iCommandPCPLC:=D2097; 
ComConveyorIO70195.i_iTaskIDPCPLC:=D2098; 
DMOV(TRUE,D2099,ComConveyorIO70195.i_diDestinationDevicePCPLC); 
ComConveyorIO70195.i_iProductIDPCPLC:=D2101;
D3090:=ComConveyorIO70195.o_iRequestPLCPC; 
D3091:=ComConveyorIO70195.o_iForceInportPLCPC;